ScreenModuleEditorView "HMI_PID_ex" 640x480
   TextField "Text field_7" at 243,29 size 43x22; Text 'вход'
      Visibility <- "Visu.view_settings"
   TextField "Text field_8" at 243,54 size 56x22; Text 'выход'
      Visibility <- "Visu.view_settings"
   IOField "I/O field_1" at 309,30 size 92x26; FormatPattern s99999.9
      Visibility <- "Visu.view_settings"
      ProcessValue <- "PIDx.Min_in"
   IOField "I/O field_2" at 309,52 size 92x26; FormatPattern s99999.9
      Visibility <- "Visu.view_settings"
      ProcessValue <- "PIDx.Min_out"
   IOField "I/O field_3" at 405,29 size 92x26; FormatPattern s99999.9
      Visibility <- "Visu.view_settings"
      ProcessValue <- "PIDx.Max_in"
   IOField "I/O field_4" at 405,51 size 92x26; FormatPattern s99999.9
      Visibility <- "Visu.view_settings"
      ProcessValue <- "PIDx.Max_out"
   Button "Button_6" at 241,105 size 68x30; TextOff 'Reset'
      on Click: SetBit("PIDx.Reset")
      Visibility <- "Visu.view_settings"
      Appearance <- "PIDx.Reset"
   IOField "I/O field_10" at 311,105 size 55x30; FormatPattern FFFF
      Visibility <- "Visu.view_settings"
      ProcessValue <- "PIDx.Warning_code"
   TextField "Text field_5" at 247,137 size 46x22; Text 'Cycle'
      Visibility <- "Visu.view_settings"
   IOField "I/O field_9" at 302,137 size 63x23; FormatPattern 99.9
      Visibility <- "Visu.view_settings"
      ProcessValue <- "PIDx.SP_Cycle"
   IOField "I/O field_15" at 368,105 size 55x30; FormatPattern FFFF
      Visibility <- "Visu.view_settings"
      ProcessValue <- "PIDx.Error_code"
      Appearance <- "PIDx.Error"
   Button "Button_2" at 426,105 size 71x30; TextOff 'Invers'
      on Click: InvertBit("PIDx.Invert")
      Visibility <- "Visu.view_settings"
      Appearance <- "PIDx.Invert"
   TextField "Text field_17" at 243,77 size 67x22; Text 'уставка'
      Visibility <- "Visu.view_settings"
   IOField "I/O field_17" at 309,75 size 92x26; FormatPattern s99999.9
      Visibility <- "Visu.view_settings"
      ProcessValue <- "PIDx.Min_SP"
   IOField "I/O field_18" at 405,74 size 92x26; FormatPattern s99999.9
      Visibility <- "Visu.view_settings"
      ProcessValue <- "PIDx.Max_SP"
   TextField "Text field_14" at 367,138 size 62x22; Text 'OnTime'
      Visibility <- "Visu.view_settings"
   IOField "I/O field_13" at 432,138 size 63x23; FormatPattern 99.9
      Visibility <- "Visu.view_settings"
      ProcessValue <- "PIDx.OnTime"
   TextField "Text field_15" at 368,168 size 65x22; Text 'OffTime'
      Visibility <- "Visu.view_settings"
   IOField "I/O field_14" at 433,168 size 63x23; FormatPattern 99.9
      Visibility <- "Visu.view_settings"
      ProcessValue <- "PIDx.OffTime"
   TextField "Text field_18" at 239,158 size 60x22; Text 'SP Low'
      Visibility <- "Visu.view_settings"
      Appearance <- "PIDx.SP_L"
   TextField "Text field_19" at 299,157 size 63x22; Text 'SP High'
      Visibility <- "Visu.view_settings"
      Appearance <- "PIDx.SP_H"
   TextField "Text field_20" at 239,182 size 56x22; Text 'In Low'
      Visibility <- "Visu.view_settings"
      Appearance <- "PIDx.In_L"
   TextField "Text field_21" at 299,181 size 59x22; Text 'In High'
      Visibility <- "Visu.view_settings"
      Appearance <- "PIDx.In_H"
   Rectangle "Rectangle_2" at 237,26 size 265x215
      Visibility <- "Visu.view_settings"
   TextField "Text field_9" at 33,59 size 15x22; Text 'K'
   TextField "Text field_10" at 33,91 size 19x22; Text 'Ti'
   IOField "I/O field_5" at 71,61 size 70x30; FormatPattern s999.99
      ProcessValue <- "PIDx.SP_P"
   IOField "I/O field_6" at 71,92 size 70x30; FormatPattern 999.9
      ProcessValue <- "PIDx.SP_Ti"
   TextField "Text field_11" at 33,124 size 23x22; Text 'Td'
   IOField "I/O field_7" at 71,123 size 70x30; FormatPattern 999.9
      ProcessValue <- "PIDx.SP_Td"
   Button "Button_4" at 73,164 size 68x30; TextOff 'Hand'
      on Click: InvertBit("PIDx.Hand")
      Appearance <- "PIDx.Hand"
   IOField "I/O field_8" at 36,201 size 109x30; FormatPattern s999.99
      ProcessValue <- "PIDx.HandValue"
   SymbolicIOField "Symbolic I/O field_1" at 147,31 size 81x24; TextOn '1'; TextOff '0'; TextList "Mode"
      ProcessValue <- "PIDx.Type"
   TextField "Text field_3" at 78,29 size 62x22; Text 'Режим:'
   TextField "Text field_12" at 155,58 size 67x22; Text 'Датчик:'
   IOField "I/O field_11" at 154,80 size 63x23; FormatPattern s999.9
      ProcessValue <- "PIDx.Value"
   TextField "Text field_13" at 149,120 size 73x22; Text 'Уставка:'
   IOField "I/O field_12" at 155,144 size 63x23; FormatPattern s999.9
      ProcessValue <- "PIDx.SP"
   IOField "I/O field_16" at 149,203 size 77x28; FormatPattern s999.9
      ProcessValue <- "PIDx.Result"
   TextField "Text field_16" at 159,181 size 53x22; Text 'Result'
   Button "Button_1" at 35,164 size 30x30; TextOff 'Text'; PictureOff "sys_volume control"
      on Click: SetBit("Visu.view_settings")
   Button "Button_3" at 241,201 size 255x30; TextOff 'Save'
      on Click: ResetBit("Visu.view_settings")
      Visibility <- "Visu.view_settings"
*)

(* ===== HMI "HMI_RT_1" =====
system functions are stored by id; their names below are inferred from use

text list "Hand": 0 'Авто'; 1 'Ручной'

graphic list "датчик1_0": 0 'Off'; 1 'On'

graphic list "Valve_hor": 1 'open'; 2 'opening'; 3 'closing'; 7 'alm_close'; 0 'close'; 4 'no_data'; 8 'alm_open'; 9 'Alarm_3'

ScreenModuleEditorView "HMI_DO_valve_hor" 1024x768
   GraphicIOField "Graphic IO Field_7" at 160,102 size 32x34; PictureList "Valve_hor"
      ProcessValue <- "Valve.Status"
   GraphicView "Graphics View" at 181,99 size 24x24; Picture "z2use"
      Visibility <- "Valve.Hand"
   Button "Button_5" at 157,94 size 48x48; TextOff 'Text'
      on Click: InvertBit("View.view_circle")
   Rectangle "Rectangle_1" at 121,21 size 112x78
      Visibility <- "View.view_circle"
   Button "Button_3" at 129,28 size 95x20; TextOff 'Авто'; TextList "Hand"
      on Click: InvertBit("Valve.Hand")
      Visibility <- "View.view_circle"
      Appearance <- "Valve.Hand"
   Button "Button_4" at 175,52 size 49x20; TextOff 'Выкл'
      on Click: ResetBit("Valve.Start_M_Fw")
      Visibility <- "View.view_circle"
   Button "Button_12" at 129,52 size 47x20; TextOff 'Вкл'
      on Click: SetBit("Valve.Start_M_Fw")
      Visibility <- "View.view_circle"
      Appearance <- "Valve.Start_M_Fw"
   TextField "Text field_1" at 129,72 size 97x22; Text 'Text'
      Visibility <- "View.view_circle"
   TextField "Text field_2" at 129,72 size 97x22; Text 'Text'
      Visibility <- "All"
*)

(* ===== HMI "HMI_RT_1" =====
system functions are stored by id; their names below are inferred from use

text list "Number": 1 'P1'; 2 'P2'; 3 'P3'; 4 'P11-A'; 5 'P12-A'; 6 'P13-A'; 7 'P14-I'; 8 'P15'; 9 'P4'; 10 'P6-A'; 11 'P7-A'; 12 'P21-A'; 13 'P22-A'; 14 'P10'; 15 'P11'; 16 'P12'; 17 'IE-P-02'; 18 'P26-I'; 19 'P27'; 20 'S27'; 21 'P24'; 22 'P25-A'; 23 'P25'; 24 'P29-A'; 25 'P31-A'; 26 'P33'; 27 'P25'; 28 'P26'; 29 'DP11'; 30 'DP12'; 31 'DP23'; 32 'DP65'

text list "Mode": 0 'Автомат'; 1 'Ручной'; 2 'Force'; 3 'Симуляция'; 4 'Удалённый'; 5 'Локальный'; 6 'Заблокирован'; 7 ''; 8 ''; 9 'Отключён'; 10 'Сервисный'

text list "Status": 0 'Выкл'; 1 'Вкл'; 2 'Остановка'; 3 'Запуск'; 4 'Авария ВЫКЛ'; 5 'Авария ВКЛ'; 6 'Авария QF'; 7 'Отключён'

text list "Hand": 0 'Авто'; 1 'Ручной'

text list "настройки": 0 'Настройки >>'; 1 'Настройки <<'

graphic list "Pump_Down": 1 'pump_ok'; 2 'pump_wait'; 3 'pump_wait_1'; 7 'down_stop'; 0 'pump_off'; 4 'pump'; 8 'down_start'; 9 'down_alm'

graphic list "Pump_Up": 1 'up_on'; 2 'up_wait'; 3 'up_wait'; 7 'up_stop'; 0 'up_off'; 4 'up_no'; 8 'up_start'; 9 'up_alm'

graphic list "Pump_Left": 1 'left_on'; 2 'left_wait'; 3 'left_wait_1'; 7 'left_stop'; 0 'left_off'; 4 'left_no'; 8 'left_start'; 9 'left_alm'

graphic list "Pump_Right": 1 'right_on'; 2 'right_wait'; 3 'right_wait_1'; 7 'right_stop'; 0 'right_off'; 4 'right_no'; 8 'right_start'; 9 'right_alm'

graphic list "V_Right": 1 'right_open_3x'; 2 'right_closing_3x'; 3 'right_opening_3x'; 7 'right_cl_alm_3xя'; 0 'right_close_3x'; 4 'right_no_3x'; 8 'right_op_alm_3x'; 9..100 'right_alm_3x'

graphic list "Z_Hor": 1 'h_open'; 2 'd_closing'; 3 'd_open'; 0 'v_close'; 4 'v_no'; 7..100 'down_alm_3x'

graphic list "Z_Vert": 1 'v_open'; 2 'd_closing_1'; 3 'd_opening'; 0 'h_close'; 4 'h_no'; 7..100 'h_alarm'

graphic list "V_Down": 1 'down_open_3x'; 2 'down_closing_3x'; 3 'down_opening_3x'; 7 'down_cl_alm_3xя'; 0 'down_close_3x'; 4 'down_no_3x'; 8 'down_op_alm_3x'; 9..100 'down_alm_3x'

graphic list "V_Up": 1 'up_open_3x'; 2 'up_closing_3x'; 3 'up_opening_3x'; 7 'up_cl_alm_3xя'; 0 'up_close_3x'; 4 'up_no_3x'; 8 'up_op_alm_3x'; 9 'up_alm_3x'

graphic list "V_Left": 1 'left_open_3x'; 2 'left_closing_3x'; 3 'left_opening_3x'; 7 'left_cl_alm_3xя'; 0 'left_close_3x'; 4 'left_no_3x'; 8 'left_op_alm_3x'; 9..100 'left_alm_3x'

ScreenModuleEditorView "HMI_M_Uni_DA" 1024x768
   Rectangle "Rectangle_3" at 452,30 size 220x193
      Visibility <- "Visu.view_settings"
   Rectangle "Rectangle_2" at 305,30 size 167x193
      Visibility <- "Visu.view_circle"
   GraphicIOField "Graphic I/O field_2" at 155,105 size 60x60; PictureList "Pump_Down"
      Visibility <- "Type"
      ProcessValue <- "M.Status"
   Button "Button_3" at 233,99 size 95x30; TextOff 'Авто'; TextList "Hand"
      on Click: InvertBit("M.Hand")
      Appearance <- "M.Hand"
      ProcessValue <- "M.Hand"
   Button "Button_4" at 279,143 size 49x30; TextOff 'Выкл'
      on Click: ResetBit("M.Start_M")
   Button "Button_7" at 341,60 size 122x20; TextOff 'Сервис'
      on Click: InvertBit("M.Trace_lock")
      Visibility <- "Visu.view_circle"
      Appearance <- "M.Trace_lock"
   Button "Button_8" at 341,87 size 122x20; TextOff 'Локально'
      on Click: InvertBit("M.Local")
      Visibility <- "Visu.view_circle"
      Appearance <- "M.Local"
   Button "Button_9" at 477,58 size 95x20; TextOff 'Force'
      on Click: InvertBit("M.Force")
      Visibility <- "Visu.view_settings"
      Appearance <- "M.Force"
   Button "Button_11" at 477,114 size 95x20; TextOff 'Simultaion'
      on Click: InvertBit("M.Sim")
      Visibility <- "Visu.view_settings"
      Appearance <- "M.Sim"
   IOField "I/O field_1" at 137,186 size 46x30; FormatPattern 999
      Visibility <- "M.Analog"
      ProcessValue <- "M.SP_A"
   IOField "I/O field_2" at 234,186 size 97x30; FormatPattern 999
      Visibility <- "M.Analog"
      ObjectEnable <- "M.Hand"
      ProcessValue <- "M.SP_M"
   Circle "Circle_4" at 650,55 size 18x18
      Visibility <- "Visu.view_settings"
      Appearance <- "M.FB_QF"
   Circle "Circle_5" at 650,83 size 18x18
      Visibility <- "Visu.view_settings"
      Appearance <- "M.FB_Run"
   TextField "Text field_4" at 580,55 size 69x18; Text 'Готовность'
      Visibility <- "Visu.view_settings"
   TextField "Text field_5" at 580,83 size 56x18; Text 'В работе'
      Visibility <- "Visu.view_settings"
   IOField "I/O field_3" at 339,136 size 28x20; FormatPattern 99
      Visibility <- "Visu.view_circle"
      ProcessValue <- "M.Wait_On_SP"
   IOField "I/O field_4" at 402,137 size 31x20; FormatPattern 99
      Visibility <- "Visu.view_circle"
      ProcessValue <- "M.Wait_Off_SP"
   TextField "Text field_6" at 344,117 size 45x18; Text 'Вкл (с)'
      Visibility <- "Visu.view_circle"
   TextField "Text field_7" at 402,117 size 53x18; Text 'Выкл (с)'
      Visibility <- "Visu.view_circle"
   Button "Button_12" at 233,143 size 47x30; TextOff 'Вкл'
      on Click: SetBit("M.Start_M")
      Appearance <- "M.Start_M"
   TextField "Text field_13" at 137,60 size 194x26; Text 'Text'
   TextField "Text field_15" at 369,159 size 64x18; Text 'Задержка:'
      Visibility <- "Visu.view_circle"
   TextField "Text field_16" at 338,179 size 36x18; Text 'пуска'
      Visibility <- "Visu.view_circle"
   IOField "I/O field_6" at 393,177 size 31x20; FormatPattern 99
      Visibility <- "Visu.view_circle"
      ProcessValue <- "M.Delay_On_SP"
   IOField "I/O field_7" at 393,200 size 30x20; FormatPattern 99
      Visibility <- "Visu.view_circle"
      ProcessValue <- "M.Delay_Off_SP"
   TextField "Text field_17" at 336,200 size 56x18; Text 'останова'
      Visibility <- "Visu.view_circle"
   IOField "I/O field_8" at 429,177 size 31x20; FormatPattern 99
      Visibility <- "Visu.view_circle"
      ProcessValue <- "M.Delay_On_Now"
   IOField "I/O field_9" at 429,200 size 30x20; FormatPattern 99
      Visibility <- "Visu.view_circle"
      ProcessValue <- "M.Delay_Off_Now"
   IOField "I/O field_10" at 367,136 size 28x20; FormatPattern 99
      Visibility <- "Visu.view_circle"
      ProcessValue <- "M.Wait_On_Now"
   IOField "I/O field_11" at 433,137 size 31x20; FormatPattern 99
      Visibility <- "Visu.view_circle"
      ProcessValue <- "M.Wait_Off_Now"
   Button "Button_16" at 477,86 size 95x20; TextOff 'Impulse'
      on Click: InvertBit("M.Impulse")
      Visibility <- "Visu.view_settings"
      Appearance <- "M.Impulse"
   Circle "Circle_1" at 650,112 size 18x18
      Visibility <- "Visu.view_settings"
      Appearance <- "M.Pos_Ok"
   Circle "Circle_2" at 650,140 size 18x18
      Visibility <- "Visu.view_settings"
      Appearance <- "M.FB_Speed_Ok"
   TextField "Text field_1" at 580,112 size 53x18; Text 'Позиция'
      Visibility <- "Visu.view_settings"
   TextField "Text field_2" at 580,140 size 57x18; Text 'Скорость'
      Visibility <- "Visu.view_settings"
   Button "Button_1" at 477,143 size 95x20; TextOff 'Analog'
      on Click: InvertBit("M.Analog")
      Visibility <- "Visu.view_settings"
      Appearance <- "M.Analog"
   Button "Button_2" at 477,171 size 61x20; TextOff 'Servo'
      on Click: InvertBit("M.Servo")
      Visibility <- "Visu.view_settings"
      Appearance <- "M.Servo"
   Button "Button_5" at 477,200 size 95x20; TextOff 'Speed'
      on Click: InvertBit("M.Speed")
      Visibility <- "Visu.view_settings"
      Appearance <- "M.Speed"
   TextField "Text field_8" at 580,160 size 36x18; Text 'Servo'
      Visibility <- "Visu.view_settings"
   IOField "I/O field_5" at 582,179 size 37x20; FormatPattern 99
      Visibility <- "Visu.view_settings"
      ProcessValue <- "M.Delay_Servo_SP"
   IOField "I/O field_12" at 582,201 size 36x20; FormatPattern 99
      Visibility <- "Visu.view_settings"
      ProcessValue <- "M.Delay_Servo_Now"
   TextField "Text field_9" at 626,159 size 40x18; Text 'Speed'
      Visibility <- "Visu.view_settings"
   IOField "I/O field_13" at 630,179 size 37x20; FormatPattern 99
      Visibility <- "Visu.view_settings"
      ProcessValue <- "M.Delay_Speed_SP"
   IOField "I/O field_14" at 630,201 size 36x20; FormatPattern 99
      Visibility <- "Visu.view_settings"
      ProcessValue <- "M.Delay_Speed_Now"
   Button "Button_6" at 137,33 size 194x22; TextOff 'Настройки >>'; TextList "настройки"
      on Click: InvertBit("Visu.view_circle"); ResetBit("Visu.view_settings")
      ProcessValue <- "Visu.view_circle"
   Button "Button_10" at 341,32 size 123x22; TextOff 'Отладка >>'
      on Click: SetBit("Visu.view_settings")
      Visibility <- "Visu.view_circle"
   Button "Button_13" at 477,32 size 192x22; TextOff 'Закрыть'
      on Click: ResetBit("Visu.view_settings")
      Visibility <- "Visu.view_settings"
   GraphicIOField "Graphic I/O field_1" at 155,105 size 60x60; PictureList "Pump_Up"
      Visibility <- "Type"
      ProcessValue <- "M.Status"
   GraphicIOField "Graphic I/O field_3" at 155,105 size 60x60; PictureList "Pump_Left"
      Visibility <- "Type"
      ProcessValue <- "M.Status"
   GraphicIOField "Graphic I/O field_4" at 155,105 size 60x60; PictureList "Pump_Right"
      Visibility <- "Type"
      ProcessValue <- "M.Status"
   IOField "I/O field_15" at 183,186 size 46x30; FormatPattern 999
      Visibility <- "M.Analog"
      ProcessValue <- "M.FB_SP"
   IOField "I/O field_16" at 537,171 size 37x20; FormatPattern 9.9
      Visibility <- "Visu.view_settings"
      ProcessValue <- "M.Servo_DB"
   GraphicIOField "Graphic I/O field_5" at 155,105 size 60x60; PictureList "V_Down"
      Visibility <- "Type"
   GraphicIOField "Graphic I/O field_6" at 155,105 size 60x60; PictureList "V_Up"
      Visibility <- "Type"
   GraphicIOField "Graphic I/O field_7" at 155,105 size 60x60; PictureList "V_Left"
      Visibility <- "Type"
   GraphicIOField "Graphic I/O field_8" at 155,105 size 60x60; PictureList "V_Right"
      Visibility <- "Type"
   GraphicIOField "Graphic I/O field_9" at 155,105 size 60x60; PictureList "Z_Hor"
      Visibility <- "Type"
   GraphicIOField "Graphic I/O field_10" at 155,105 size 60x60; PictureList "Z_Vert"
      Visibility <- "Type"
   GraphicView "Graphic view_1" at 134,87 size 30x30; Picture "z2use_3"
      Visibility <- "M.Hand"
   GraphicView "Graphic view_8" at 204,86 size 30x30; Picture "force"
      Visibility <- "M.Force"
   GraphicView "Graphic view_10" at 133,128 size 50x54; Picture "lock_32x32"
      Visibility <- "M.Lock"
   GraphicView "Graphic view_11" at 192,146 size 30x30; Picture "service"
      Visibility <- "M.Trace_lock"
   GraphicView "Graphic view_12" at 168,86 size 30x30; Picture "local"
      Visibility <- "M.Local"
*)

(* ===== HMI "HMI_RT_1" =====
system functions are stored by id; their names below are inferred from use

text list "Number": 1 'P1'; 2 'P2'; 3 'P3'; 4 'P11-A'; 5 'P12-A'; 6 'P13-A'; 7 'P14-I'; 8 'P15'; 9 'P4'; 10 'P6-A'; 11 'P7-A'; 12 'P21-A'; 13 'P22-A'; 14 'P10'; 15 'P11'; 16 'P12'; 17 'IE-P-02'; 18 'P26-I'; 19 'P27'; 20 'S27'; 21 'P24'; 22 'P25-A'; 23 'P25'; 24 'P29-A'; 25 'P31-A'; 26 'P33'; 27 'P25'; 28 'P26'; 29 'DP11'; 30 'DP12'; 31 'DP23'; 32 'DP65'

text list "Mode": 0 'Автомат'; 1 'Ручной'; 2 'Force'; 3 'Симуляция'; 4 'Удалённый'; 5 'Локальный'; 6 'Заблокирован'; 7 ''; 8 ''; 9 'Отключён'; 10 'Сервисный'

text list "Status": 0 'Выкл'; 1 'Вкл'; 2 'Остановка'; 3 'Запуск'; 4 'Авария ВЫКЛ'; 5 'Авария ВКЛ'; 6 'Авария QF'; 7 'Отключён'

text list "Hand": 0 'Авто'; 1 'Ручной'

text list "настройки": 0 'Настройки >>'; 1 'Настройки <<'

graphic list "Pump_Down": 1 'pump_ok'; 2 'pump_wait'; 3 'pump_wait_1'; 7 'down_stop'; 0 'pump_off'; 4 'pump'; 8 'down_start'; 9 'down_alm'

graphic list "Pump_Up": 1 'up_on'; 2 'up_wait'; 3 'up_wait'; 7 'up_stop'; 0 'up_off'; 4 'up_no'; 8 'up_start'; 9 'up_alm'

graphic list "Pump_Left": 1 'left_on'; 2 'left_wait'; 3 'left_wait_1'; 7 'left_stop'; 0 'left_off'; 4 'left_no'; 8 'left_start'; 9 'left_alm'

graphic list "Pump_Right": 1 'right_on'; 2 'right_wait'; 3 'right_wait_1'; 7 'right_stop'; 0 'right_off'; 4 'right_no'; 8 'right_start'; 9 'right_alm'

graphic list "V_Right": 1 'right_open_3x'; 2 'right_closing_3x'; 3 'right_opening_3x'; 7 'right_cl_alm_3xя'; 0 'right_close_3x'; 4 'right_no_3x'; 8 'right_op_alm_3x'; 9..100 'right_alm_3x'

graphic list "Z_Hor": 1 'h_open'; 2 'd_closing'; 3 'd_open'; 0 'v_close'; 4 'v_no'; 7..100 'down_alm_3x'

graphic list "Z_Vert": 1 'v_open'; 2 'd_closing_1'; 3 'd_opening'; 0 'h_close'; 4 'h_no'; 7..100 'h_alarm'

graphic list "V_Down": 1 'down_open_3x'; 2 'down_closing_3x'; 3 'down_opening_3x'; 7 'down_cl_alm_3xя'; 0 'down_close_3x'; 4 'down_no_3x'; 8 'down_op_alm_3x'; 9..100 'down_alm_3x'

graphic list "V_Up": 1 'up_open_3x'; 2 'up_closing_3x'; 3 'up_opening_3x'; 7 'up_cl_alm_3xя'; 0 'up_close_3x'; 4 'up_no_3x'; 8 'up_op_alm_3x'; 9 'up_alm_3x'

graphic list "V_Left": 1 'left_open_3x'; 2 'left_closing_3x'; 3 'left_opening_3x'; 7 'left_cl_alm_3xя'; 0 'left_close_3x'; 4 'left_no_3x'; 8 'left_op_alm_3x'; 9..100 'left_alm_3x'

ScreenModuleEditorView "HMI_M_Uni_DA" 1024x768
   Rectangle "Rectangle_3" at 452,30 size 168x194
      Visibility <- "Visu.view_settings"
   Rectangle "Rectangle_2" at 305,30 size 150x194
      Visibility <- "Visu.view_circle"
   GraphicIOField "Graphic I/O field_2" at 161,105 size 60x60; PictureList "Pump_Down"
      Visibility <- "Type"
      ProcessValue <- "M.Status"
   Button "Button_3" at 233,99 size 90x30; TextOff 'Авто'; TextList "Hand"
      on Click: InvertBit("M.Hand")
      ProcessValue <- "M.Hand"
      Appearance <- "M.Hand"
   Button "Button_4" at 277,143 size 45x30; TextOff 'Выкл'
      on Click: ResetBit("M.Start_M")
   Button "Button_7" at 329,60 size 122x20; TextOff 'Сервис'
      on Click: InvertBit("M.Trace_lock")
      Visibility <- "Visu.view_circle"
      Appearance <- "M.Trace_lock"
   Button "Button_8" at 329,87 size 122x20; TextOff 'Локально'
      on Click: InvertBit("M.Local")
      Visibility <- "Visu.view_circle"
      Appearance <- "M.Local"
   Button "Button_9" at 461,58 size 70x20; TextOff 'Force'
      on Click: InvertBit("M.Force")
      Visibility <- "Visu.view_settings"
      Appearance <- "M.Force"
   Button "Button_11" at 461,114 size 70x20; TextOff 'Sim'
      on Click: InvertBit("M.Sim")
      Visibility <- "Visu.view_settings"
      Appearance <- "M.Sim"
   IOField "I/O field_1" at 148,186 size 46x30; FormatPattern 999
      Visibility <- "M.Analog"
      ProcessValue <- "M.SP_A"
   IOField "I/O field_2" at 250,186 size 73x30; FormatPattern 999
      Visibility <- "M.Analog"
      ObjectEnable <- "M.Hand"
      ProcessValue <- "M.SP_M"
   Circle "Circle_4" at 598,55 size 18x18
      Visibility <- "Visu.view_settings"
      Appearance <- "M.FB_QF"
   Circle "Circle_5" at 598,83 size 18x18
      Visibility <- "Visu.view_settings"
      Appearance <- "M.FB_Run"
   TextField "Text field_4" at 535,55 size 37x18; Text 'Готов'
      Visibility <- "Visu.view_settings"
   TextField "Text field_5" at 535,83 size 56x18; Text 'В работе'
      Visibility <- "Visu.view_settings"
   IOField "I/O field_3" at 327,137 size 30x20; FormatPattern 99
      Visibility <- "Visu.view_circle"
      ProcessValue <- "M.Wait_On_SP"
   IOField "I/O field_4" at 389,137 size 30x20; FormatPattern 99
      Visibility <- "Visu.view_circle"
      ProcessValue <- "M.Wait_Off_SP"
   TextField "Text field_6" at 332,117 size 45x18; Text 'Вкл (с)'
      Visibility <- "Visu.view_circle"
   TextField "Text field_7" at 390,117 size 53x18; Text 'Выкл (с)'
      Visibility <- "Visu.view_circle"
   Button "Button_12" at 233,143 size 45x30; TextOff 'Вкл'
      on Click: SetBit("M.Start_M")
      Appearance <- "M.Start_M"
   TextField "Text field_13" at 147,60 size 177x26; Text 'Text'
   TextField "Text field_15" at 357,159 size 64x18; Text 'Задержка:'
      Visibility <- "Visu.view_circle"
   TextField "Text field_16" at 326,179 size 36x18; Text 'пуска'
      Visibility <- "Visu.view_circle"
   IOField "I/O field_6" at 381,177 size 30x20; FormatPattern 99
      Visibility <- "Visu.view_circle"
      ProcessValue <- "M.Delay_On_SP"
   IOField "I/O field_7" at 381,200 size 30x20; FormatPattern 99
      Visibility <- "Visu.view_circle"
      ProcessValue <- "M.Delay_Off_SP"
   TextField "Text field_17" at 324,200 size 56x18; Text 'останова'
      Visibility <- "Visu.view_circle"
   IOField "I/O field_8" at 411,177 size 30x20; FormatPattern 99
      Visibility <- "Visu.view_circle"
      ProcessValue <- "M.Delay_On_Now"
   IOField "I/O field_9" at 411,200 size 30x20; FormatPattern 99
      Visibility <- "Visu.view_circle"
      ProcessValue <- "M.Delay_Off_Now"
   IOField "I/O field_10" at 356,137 size 30x20; FormatPattern 99
      Visibility <- "Visu.view_circle"
      ProcessValue <- "M.Wait_On_Now"
   IOField "I/O field_11" at 419,137 size 30x20; FormatPattern 99
      Visibility <- "Visu.view_circle"
      ProcessValue <- "M.Wait_Off_Now"
   Button "Button_16" at 461,86 size 70x20; TextOff 'Impulse'
      on Click: InvertBit("M.Impulse")
      Visibility <- "Visu.view_settings"
      Appearance <- "M.Impulse"
   Circle "Circle_1" at 598,112 size 18x18
      Visibility <- "Visu.view_settings"
      Appearance <- "M.Pos_Ok"
   Circle "Circle_2" at 598,140 size 18x18
      Visibility <- "Visu.view_settings"
      Appearance <- "M.FB_Speed_Ok"
   TextField "Text field_1" at 535,112 size 53x18; Text 'Позиция'
      Visibility <- "Visu.view_settings"
   TextField "Text field_2" at 535,140 size 57x18; Text 'Скорость'
      Visibility <- "Visu.view_settings"
   Button "Button_1" at 461,143 size 70x20; TextOff 'Analog'
      on Click: InvertBit("M.Analog")
      Visibility <- "Visu.view_settings"
      Appearance <- "M.Analog"
   Button "Button_2" at 461,171 size 50x20; TextOff 'Servo'
      on Click: InvertBit("M.Servo")
      Visibility <- "Visu.view_settings"
      Appearance <- "M.Servo"
   Button "Button_5" at 461,200 size 70x20; TextOff 'Speed'
      on Click: InvertBit("M.Speed")
      Visibility <- "Visu.view_settings"
      Appearance <- "M.Speed"
   TextField "Text field_8" at 539,160 size 36x18; Text 'Servo'
      Visibility <- "Visu.view_settings"
   IOField "I/O field_5" at 541,179 size 35x20; FormatPattern 99
      Visibility <- "Visu.view_settings"
      ProcessValue <- "M.Delay_Servo_SP"
   IOField "I/O field_12" at 541,201 size 35x20; FormatPattern 99
      Visibility <- "Visu.view_settings"
      ProcessValue <- "M.Delay_Servo_Now"
   TextField "Text field_9" at 576,159 size 40x18; Text 'Speed'
      Visibility <- "Visu.view_settings"
   IOField "I/O field_13" at 581,179 size 35x20; FormatPattern 99
      Visibility <- "Visu.view_settings"
      ProcessValue <- "M.Delay_Speed_SP"
   IOField "I/O field_14" at 581,201 size 35x20; FormatPattern 99
      Visibility <- "Visu.view_settings"
      ProcessValue <- "M.Delay_Speed_Now"
   Button "Button_6" at 147,33 size 178x22; TextOff 'Настройки >>'; TextList "настройки"
      on Click: InvertBit("Visu.view_circle"); ResetBit("Visu.view_settings")
      ProcessValue <- "Visu.view_circle"
   Button "Button_10" at 329,33 size 123x22; TextOff 'Отладка >>'
      on Click: SetBit("Visu.view_settings")
      Visibility <- "Visu.view_circle"
   Button "Button_13" at 461,33 size 156x22; TextOff 'Закрыть'
      on Click: ResetBit("Visu.view_settings")
      Visibility <- "Visu.view_settings"
   GraphicIOField "Graphic I/O field_1" at 161,105 size 60x60; PictureList "Pump_Up"
      Visibility <- "Type"
      ProcessValue <- "M.Status"
   GraphicIOField "Graphic I/O field_3" at 161,105 size 60x60; PictureList "Pump_Left"
      Visibility <- "Type"
      ProcessValue <- "M.Status"
   GraphicIOField "Graphic I/O field_4" at 161,105 size 60x60; PictureList "Pump_Right"
      Visibility <- "Type"
      ProcessValue <- "M.Status"
   IOField "I/O field_15" at 194,186 size 46x30; FormatPattern 999
      Visibility <- "M.Analog"
      ProcessValue <- "M.FB_SP"
   IOField "I/O field_16" at 511,171 size 28x20; FormatPattern 9.9
      Visibility <- "Visu.view_settings"
      ProcessValue <- "M.Servo_DB"
   GraphicIOField "Graphic I/O field_5" at 161,105 size 60x60; PictureList "V_Down"
      Visibility <- "Type"
   GraphicIOField "Graphic I/O field_6" at 161,105 size 60x60; PictureList "V_Up"
      Visibility <- "Type"
   GraphicIOField "Graphic I/O field_7" at 161,105 size 60x60; PictureList "V_Left"
      Visibility <- "Type"
   GraphicIOField "Graphic I/O field_8" at 161,105 size 60x60; PictureList "V_Right"
      Visibility <- "Type"
   GraphicIOField "Graphic I/O field_9" at 161,105 size 60x60; PictureList "Z_Hor"
      Visibility <- "Type"
   GraphicIOField "Graphic I/O field_10" at 161,105 size 60x60; PictureList "Z_Vert"
      Visibility <- "Type"
   GraphicView "Graphic view_1" at 149,87 size 30x30; Picture "z2use_3"
      Visibility <- "M.Hand"
   GraphicView "Graphic view_8" at 207,86 size 30x30; Picture "force"
      Visibility <- "M.Force"
   GraphicView "Graphic view_10" at 143,128 size 50x54; Picture "lock_32x32"
      Visibility <- "M.Lock"
   GraphicView "Graphic view_11" at 199,146 size 30x30; Picture "service"
      Visibility <- "M.Trace_lock"
   GraphicView "Graphic view_12" at 179,86 size 30x30; Picture "local"
      Visibility <- "M.Local"
*)

(* ===== HMI "HMI_RT_1" =====
system functions are stored by id; their names below are inferred from use

text list "Number": 1 'P1'; 2 'P2'; 3 'P3'; 4 'P11-A'; 5 'P12-A'; 6 'P13-A'; 7 'P14-I'; 8 'P15'; 9 'P4'; 10 'P6-A'; 11 'P7-A'; 12 'P21-A'; 13 'P22-A'; 14 'P10'; 15 'P11'; 16 'P12'; 17 'IE-P-02'; 18 'P26-I'; 19 'P27'; 20 'S27'; 21 'P24'; 22 'P25-A'; 23 'P25'; 24 'P29-A'; 25 'P31-A'; 26 'P33'; 27 'P25'; 28 'P26'; 29 'DP11'; 30 'DP12'; 31 'DP23'; 32 'DP65'

text list "Mode": 0 'Автомат'; 1 'Ручной'; 2 'Force'; 3 'Симуляция'; 4 'Удалённый'; 5 'Локальный'; 6 'Заблокирован'; 7 ''; 8 ''; 9 'Отключён'; 10 'Сервисный'

text list "Status": 0 'Выкл'; 1 'Вкл'; 2 'Остановка'; 3 'Запуск'; 4 'Авария ВЫКЛ'; 5 'Авария ВКЛ'; 6 'Авария QF'; 7 'Отключён'

text list "Hand": 0 'Авто'; 1 'Ручной'

graphic list "Start_M": 0 'off'; 1 'on_2'

graphic list "Pump_Down": 1 'pump_ok'; 2 'pump_wait'; 3 'pump_wait_1'; 7 'down_stop'; 0 'pump_off'; 4 'pump'; 8 'down_start'; 9 'down_alm'

graphic list "Pump_Left": 1 'left_on'; 2 'left_wait'; 3 'left_wait_1'; 7 'left_stop'; 0 'left_off'; 4 'left_no'; 8 'left_start'; 9 'left_alm'

graphic list "Pump_Right": 1 'right_on'; 2 'right_wait'; 3 'right_wait_1'; 7 'right_stop'; 0 'right_off'; 4 'right_no'; 8 'right_start'; 9 'right_alm'

graphic list "Pump_Up": 1 'up_on'; 2 'up_wait'; 3 'up_wait'; 7 'up_stop'; 0 'up_off'; 4 'up_no'; 8 'up_start'; 9 'up_alm'

graphic list "V_Down": 1 'down_open_3x'; 2 'down_closing_3x'; 3 'down_opening_3x'; 7 'down_cl_alm_3xя'; 0 'down_close_3x'; 4 'down_no_3x'; 8 'down_op_alm_3x'; 9..100 'down_alm_3x'

graphic list "V_Left": 1 'left_open_3x'; 2 'left_closing_3x'; 3 'left_opening_3x'; 7 'left_cl_alm_3xя'; 0 'left_close_3x'; 4 'left_no_3x'; 8 'left_op_alm_3x'; 9..100 'left_alm_3x'

graphic list "V_Right": 1 'right_open_3x'; 2 'right_closing_3x'; 3 'right_opening_3x'; 7 'right_cl_alm_3xя'; 0 'right_close_3x'; 4 'right_no_3x'; 8 'right_op_alm_3x'; 9..100 'right_alm_3x'

graphic list "V_Up": 1 'up_open_3x'; 2 'up_closing_3x'; 3 'up_opening_3x'; 7 'up_cl_alm_3xя'; 0 'up_close_3x'; 4 'up_no_3x'; 8 'up_op_alm_3x'; 9 'up_alm_3x'

graphic list "Z_Hor": 1 'h_open'; 2 'd_closing'; 3 'd_opening_1'; 0 'v_close'; 4 'v_no'; 7..100 'down_alm_3x'

graphic list "Z_Vert": 1 'v_open'; 2 'd_closing_1'; 3 'd_opening'; 0 'h_close'; 4 'h_no'; 7..100 'h_alarm'